(* Logix 5000 project; controller MV vendor 1 type 14 code 217 rev 31.11; software revision 31.00; part 22 of 53 *)
(* tags used below, declared in another part *)
   CheckTimeMask : INT;
   CWD : CHECKWORD_FLAGS;
   Delphi_Does_Eng_Func : BOOL;
   MC_CD_T1 : PlantItem;   // CD_T1
   MC_CD_T2 : PlantItem;   // CD_T2
   MC_CH2_LF1 : PlantItem;   // CH2_LF1
   MC_FL_D1 : PlantItem;   // FL_D1
   MC_FL_D2 : PlantItem;   // FL_D2
   MC_FL_PR : PlantItem;   // FL_PR
   MC_N255 : INT[255];   // CHECKWORDS Plant item checkword s
   MC_SPV1 : PlantItem;   // SPV1
   MC_SPV2 : PlantItem;   // SPV2
   MC_SPV3 : PlantItem;   // SPV3
   MC_SPV4 : PlantItem;   // SPV4
   MC_SPV5 : PlantItem;   // SPV5
   MC_SV1 : PlantItem;   // SV1
   MC_SV2 : PlantItem;   // SV2
   TempChecktime : DINT;
(* MC_Common, continued *)

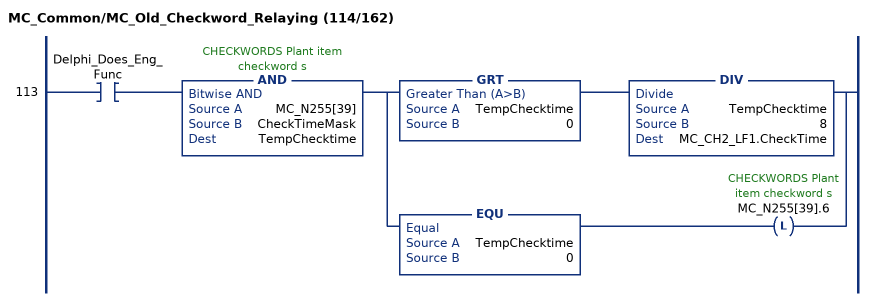
   [picture p386: MC_Common/MC_Old_Checkword_Relaying rungs 113-113]
   113: XIC(Delphi_Does_Eng_Func)AND(MC_N255[39],CheckTimeMask,TempChecktime)[GRT(TempChecktime,0) DIV(TempChecktime,8,MC_CH2_LF1.CheckTime) ,EQU(TempChecktime,0) OTL(MC_N255[39].6) ];
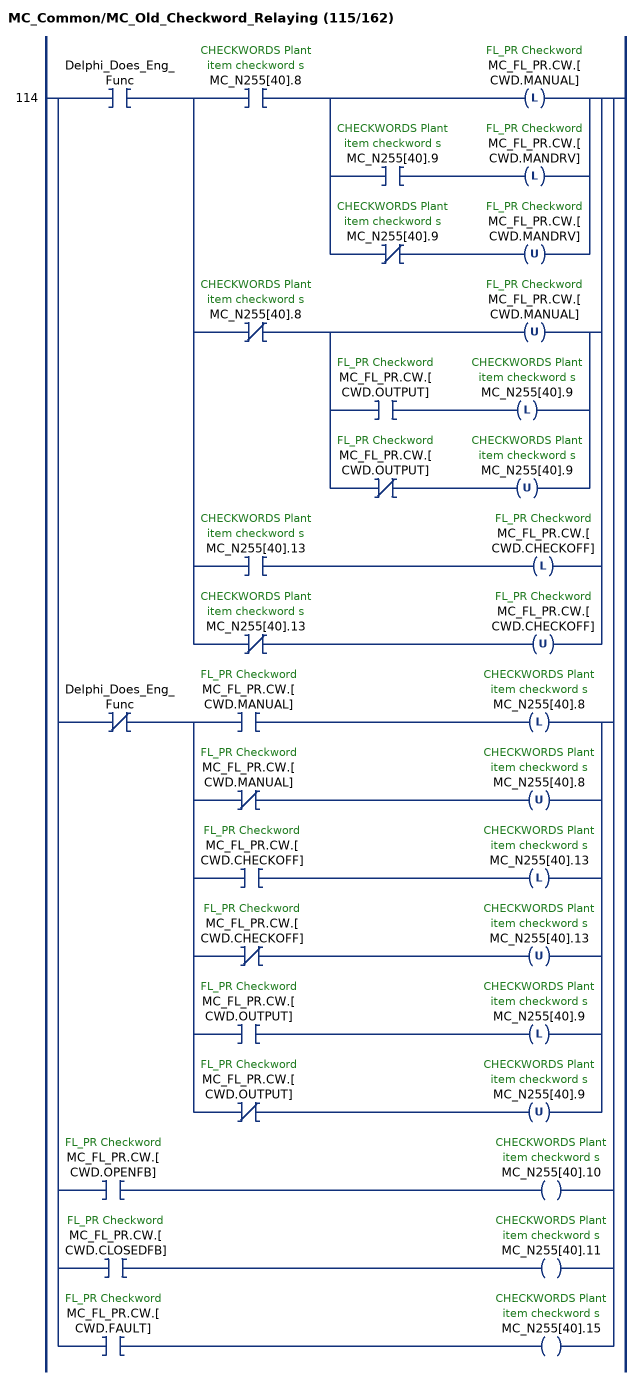
   114: [XIC(Delphi_Does_Eng_Func) [[XIC(MC_N255[40].8) [OTL(MC_FL_PR.CW.[CWD.MANUAL]) ,XIC(MC_N255[40].9) OTL(MC_FL_PR.CW.[CWD.MANDRV]) ,XIO(MC_N255[40].9) OTU(MC_FL_PR.CW.[CWD.MANDRV]) ] ,XIO(MC_N255[40].8) [OTU(MC_FL_PR.CW.[CWD.MANUAL]) ,[XIC(MC_FL_PR.CW.[CWD.OUTPUT]) OTL(MC_N255[40].9) ,XIO(MC_FL_PR.CW.[CWD.OUTPUT]) OTU(MC_N255[40].9) ] ] ] ,[XIC(MC_N255[40].13) OTL(MC_FL_PR.CW.[CWD.CHECKOFF]) ,XIO(MC_N255[40].13) OTU(MC_FL_PR.CW.[CWD.CHECKOFF]) ] ] ,XIO(Delphi_Does_Eng_Func) [[XIC(MC_FL_PR.CW.[CWD.MANUAL]) OTL(MC_N255[40].8) ,XIO(MC_FL_PR.CW.[CWD.MANUAL]) OTU(MC_N255[40].8) ] ,[XIC(MC_FL_PR.CW.[CWD.CHECKOFF]) OTL(MC_N255[40].13) ,XIO(MC_FL_PR.CW.[CWD.CHECKOFF]) OTU(MC_N255[40].13) ] ,[XIC(MC_FL_PR.CW.[CWD.OUTPUT]) OTL(MC_N255[40].9) ,XIO(MC_FL_PR.CW.[CWD.OUTPUT]) OTU(MC_N255[40].9) ] ] ,XIC(MC_FL_PR.CW.[CWD.OPENFB]) OTE(MC_N255[40].10) ,XIC(MC_FL_PR.CW.[CWD.CLOSEDFB]) OTE(MC_N255[40].11) ,XIC(MC_FL_PR.CW.[CWD.FAULT]) OTE(MC_N255[40].15) ];
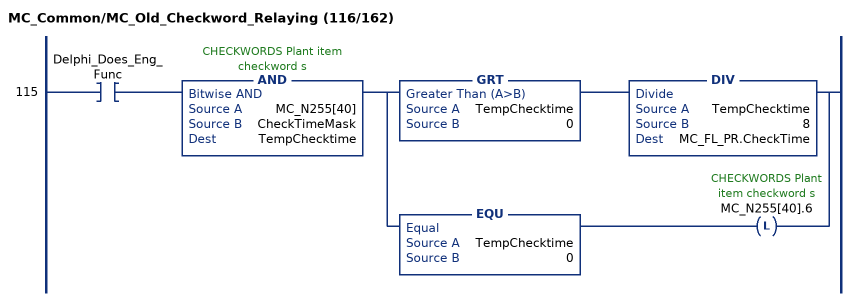
   115: XIC(Delphi_Does_Eng_Func)AND(MC_N255[40],CheckTimeMask,TempChecktime)[GRT(TempChecktime,0) DIV(TempChecktime,8,MC_FL_PR.CheckTime) ,EQU(TempChecktime,0) OTL(MC_N255[40].6) ];
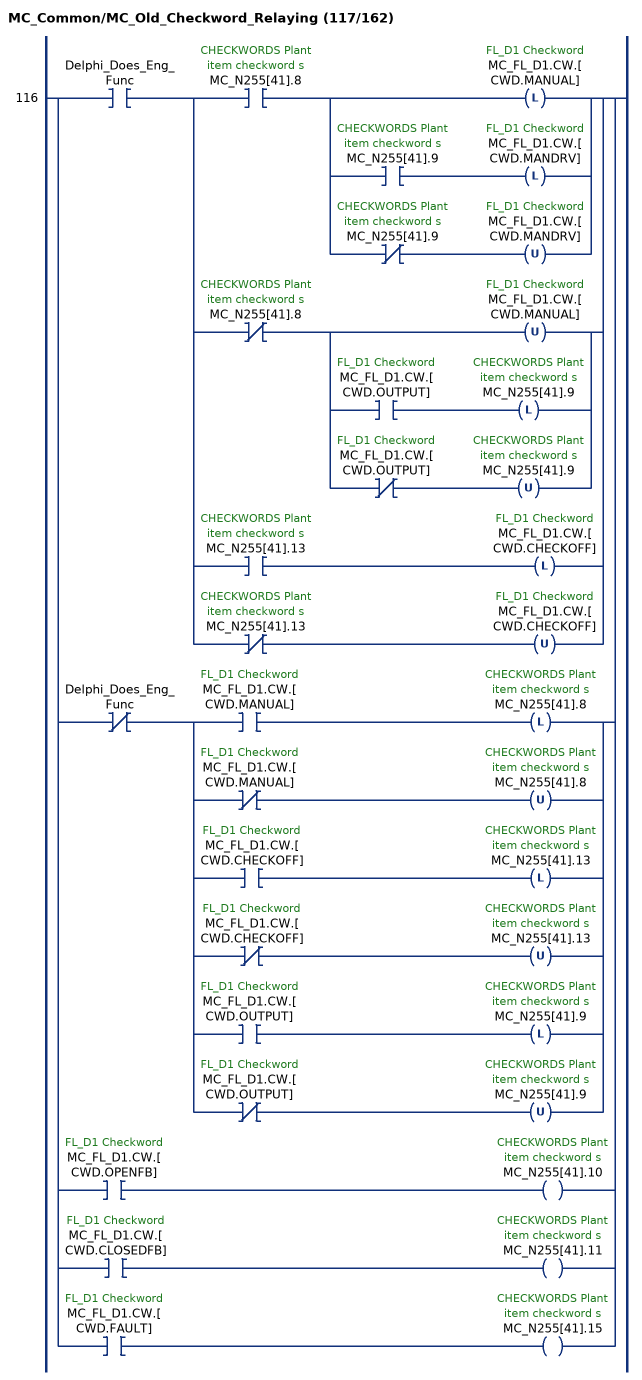
   116: [XIC(Delphi_Does_Eng_Func) [[XIC(MC_N255[41].8) [OTL(MC_FL_D1.CW.[CWD.MANUAL]) ,XIC(MC_N255[41].9) OTL(MC_FL_D1.CW.[CWD.MANDRV]) ,XIO(MC_N255[41].9) OTU(MC_FL_D1.CW.[CWD.MANDRV]) ] ,XIO(MC_N255[41].8) [OTU(MC_FL_D1.CW.[CWD.MANUAL]) ,[XIC(MC_FL_D1.CW.[CWD.OUTPUT]) OTL(MC_N255[41].9) ,XIO(MC_FL_D1.CW.[CWD.OUTPUT]) OTU(MC_N255[41].9) ] ] ] ,[XIC(MC_N255[41].13) OTL(MC_FL_D1.CW.[CWD.CHECKOFF]) ,XIO(MC_N255[41].13) OTU(MC_FL_D1.CW.[CWD.CHECKOFF]) ] ] ,XIO(Delphi_Does_Eng_Func) [[XIC(MC_FL_D1.CW.[CWD.MANUAL]) OTL(MC_N255[41].8) ,XIO(MC_FL_D1.CW.[CWD.MANUAL]) OTU(MC_N255[41].8) ] ,[XIC(MC_FL_D1.CW.[CWD.CHECKOFF]) OTL(MC_N255[41].13) ,XIO(MC_FL_D1.CW.[CWD.CHECKOFF]) OTU(MC_N255[41].13) ] ,[XIC(MC_FL_D1.CW.[CWD.OUTPUT]) OTL(MC_N255[41].9) ,XIO(MC_FL_D1.CW.[CWD.OUTPUT]) OTU(MC_N255[41].9) ] ] ,XIC(MC_FL_D1.CW.[CWD.OPENFB]) OTE(MC_N255[41].10) ,XIC(MC_FL_D1.CW.[CWD.CLOSEDFB]) OTE(MC_N255[41].11) ,XIC(MC_FL_D1.CW.[CWD.FAULT]) OTE(MC_N255[41].15) ];
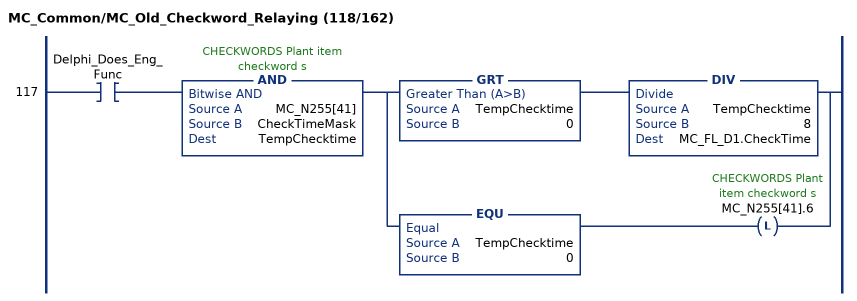
   117: XIC(Delphi_Does_Eng_Func)AND(MC_N255[41],CheckTimeMask,TempChecktime)[GRT(TempChecktime,0) DIV(TempChecktime,8,MC_FL_D1.CheckTime) ,EQU(TempChecktime,0) OTL(MC_N255[41].6) ];
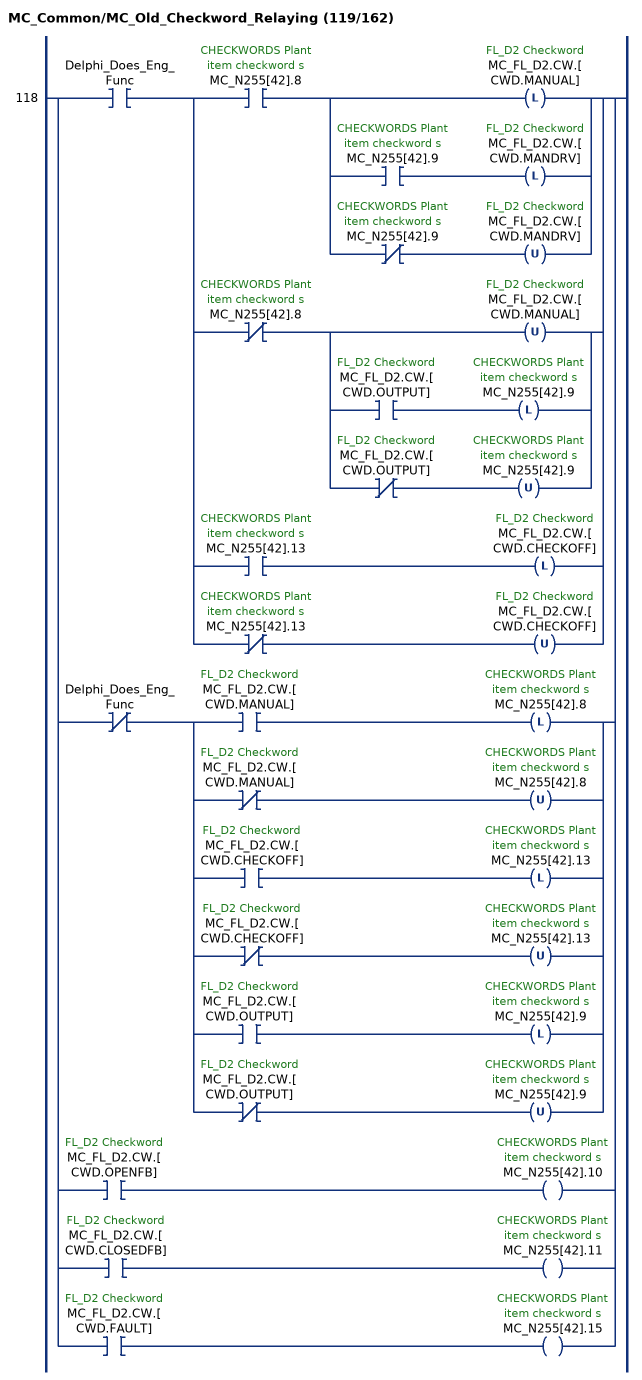
   118: [XIC(Delphi_Does_Eng_Func) [[XIC(MC_N255[42].8) [OTL(MC_FL_D2.CW.[CWD.MANUAL]) ,XIC(MC_N255[42].9) OTL(MC_FL_D2.CW.[CWD.MANDRV]) ,XIO(MC_N255[42].9) OTU(MC_FL_D2.CW.[CWD.MANDRV]) ] ,XIO(MC_N255[42].8) [OTU(MC_FL_D2.CW.[CWD.MANUAL]) ,[XIC(MC_FL_D2.CW.[CWD.OUTPUT]) OTL(MC_N255[42].9) ,XIO(MC_FL_D2.CW.[CWD.OUTPUT]) OTU(MC_N255[42].9) ] ] ] ,[XIC(MC_N255[42].13) OTL(MC_FL_D2.CW.[CWD.CHECKOFF]) ,XIO(MC_N255[42].13) OTU(MC_FL_D2.CW.[CWD.CHECKOFF]) ] ] ,XIO(Delphi_Does_Eng_Func) [[XIC(MC_FL_D2.CW.[CWD.MANUAL]) OTL(MC_N255[42].8) ,XIO(MC_FL_D2.CW.[CWD.MANUAL]) OTU(MC_N255[42].8) ] ,[XIC(MC_FL_D2.CW.[CWD.CHECKOFF]) OTL(MC_N255[42].13) ,XIO(MC_FL_D2.CW.[CWD.CHECKOFF]) OTU(MC_N255[42].13) ] ,[XIC(MC_FL_D2.CW.[CWD.OUTPUT]) OTL(MC_N255[42].9) ,XIO(MC_FL_D2.CW.[CWD.OUTPUT]) OTU(MC_N255[42].9) ] ] ,XIC(MC_FL_D2.CW.[CWD.OPENFB]) OTE(MC_N255[42].10) ,XIC(MC_FL_D2.CW.[CWD.CLOSEDFB]) OTE(MC_N255[42].11) ,XIC(MC_FL_D2.CW.[CWD.FAULT]) OTE(MC_N255[42].15) ];
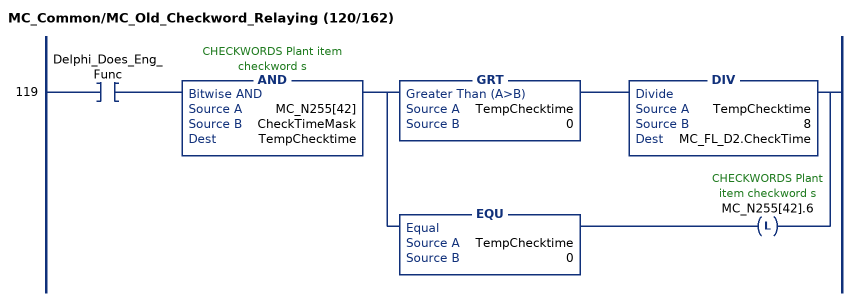
   119: XIC(Delphi_Does_Eng_Func)AND(MC_N255[42],CheckTimeMask,TempChecktime)[GRT(TempChecktime,0) DIV(TempChecktime,8,MC_FL_D2.CheckTime) ,EQU(TempChecktime,0) OTL(MC_N255[42].6) ];
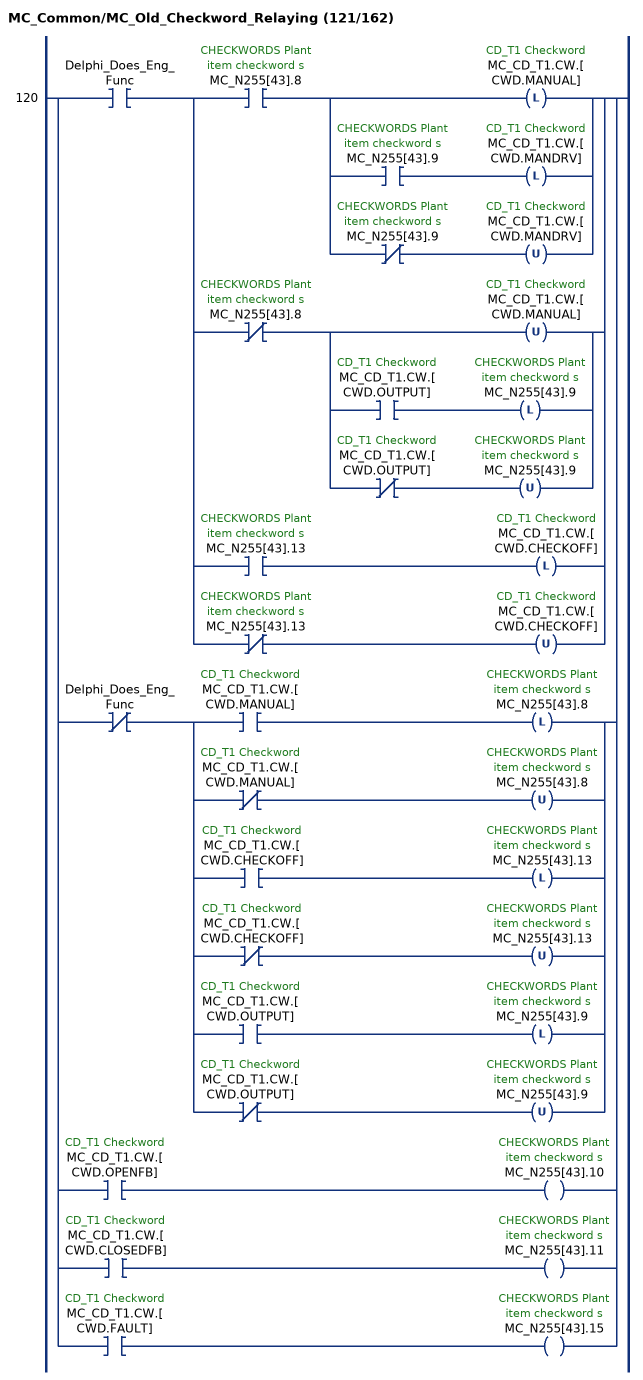
   120: [XIC(Delphi_Does_Eng_Func) [[XIC(MC_N255[43].8) [OTL(MC_CD_T1.CW.[CWD.MANUAL]) ,XIC(MC_N255[43].9) OTL(MC_CD_T1.CW.[CWD.MANDRV]) ,XIO(MC_N255[43].9) OTU(MC_CD_T1.CW.[CWD.MANDRV]) ] ,XIO(MC_N255[43].8) [OTU(MC_CD_T1.CW.[CWD.MANUAL]) ,[XIC(MC_CD_T1.CW.[CWD.OUTPUT]) OTL(MC_N255[43].9) ,XIO(MC_CD_T1.CW.[CWD.OUTPUT]) OTU(MC_N255[43].9) ] ] ] ,[XIC(MC_N255[43].13) OTL(MC_CD_T1.CW.[CWD.CHECKOFF]) ,XIO(MC_N255[43].13) OTU(MC_CD_T1.CW.[CWD.CHECKOFF]) ] ] ,XIO(Delphi_Does_Eng_Func) [[XIC(MC_CD_T1.CW.[CWD.MANUAL]) OTL(MC_N255[43].8) ,XIO(MC_CD_T1.CW.[CWD.MANUAL]) OTU(MC_N255[43].8) ] ,[XIC(MC_CD_T1.CW.[CWD.CHECKOFF]) OTL(MC_N255[43].13) ,XIO(MC_CD_T1.CW.[CWD.CHECKOFF]) OTU(MC_N255[43].13) ] ,[XIC(MC_CD_T1.CW.[CWD.OUTPUT]) OTL(MC_N255[43].9) ,XIO(MC_CD_T1.CW.[CWD.OUTPUT]) OTU(MC_N255[43].9) ] ] ,XIC(MC_CD_T1.CW.[CWD.OPENFB]) OTE(MC_N255[43].10) ,XIC(MC_CD_T1.CW.[CWD.CLOSEDFB]) OTE(MC_N255[43].11) ,XIC(MC_CD_T1.CW.[CWD.FAULT]) OTE(MC_N255[43].15) ];
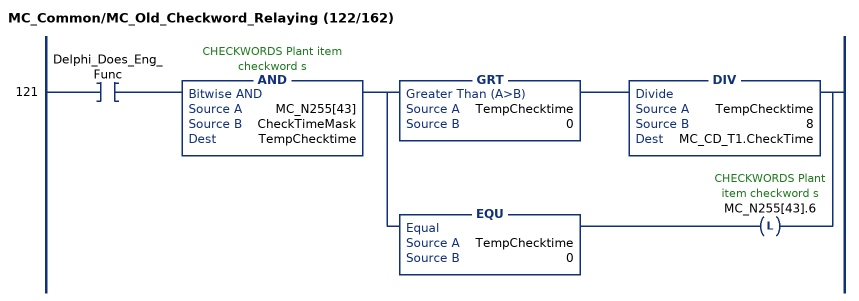
   121: XIC(Delphi_Does_Eng_Func)AND(MC_N255[43],CheckTimeMask,TempChecktime)[GRT(TempChecktime,0) DIV(TempChecktime,8,MC_CD_T1.CheckTime) ,EQU(TempChecktime,0) OTL(MC_N255[43].6) ];
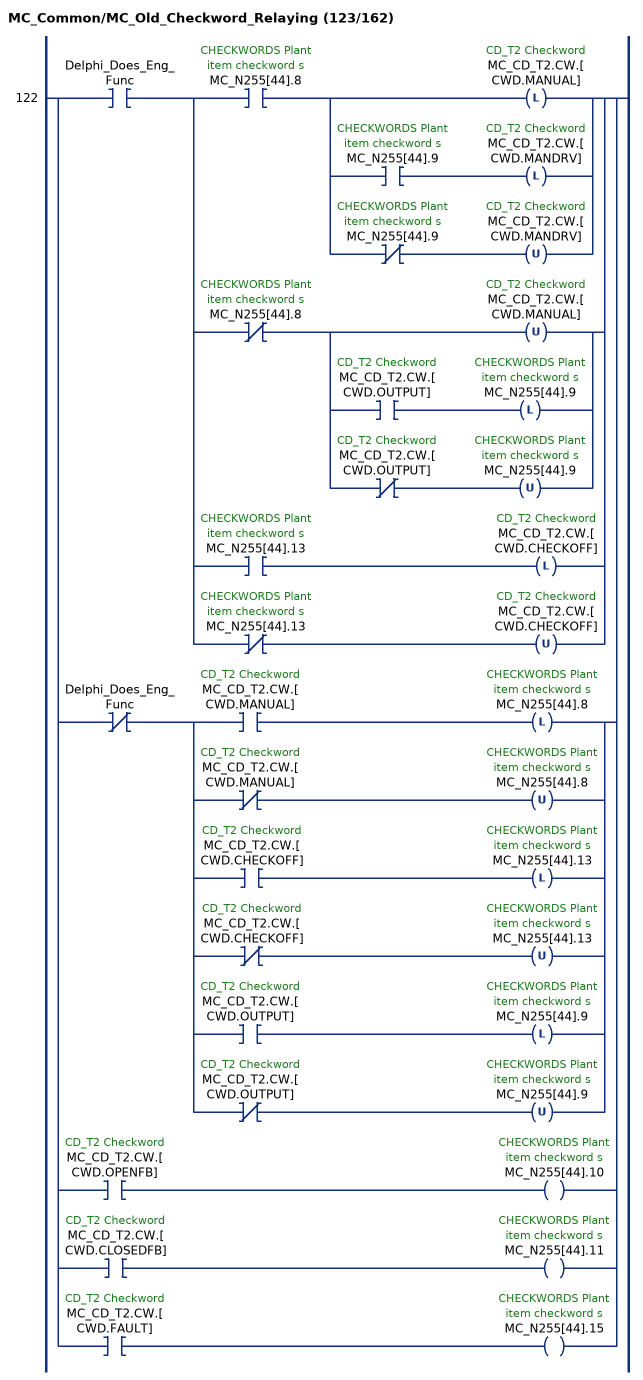
   122: [XIC(Delphi_Does_Eng_Func) [[XIC(MC_N255[44].8) [OTL(MC_CD_T2.CW.[CWD.MANUAL]) ,XIC(MC_N255[44].9) OTL(MC_CD_T2.CW.[CWD.MANDRV]) ,XIO(MC_N255[44].9) OTU(MC_CD_T2.CW.[CWD.MANDRV]) ] ,XIO(MC_N255[44].8) [OTU(MC_CD_T2.CW.[CWD.MANUAL]) ,[XIC(MC_CD_T2.CW.[CWD.OUTPUT]) OTL(MC_N255[44].9) ,XIO(MC_CD_T2.CW.[CWD.OUTPUT]) OTU(MC_N255[44].9) ] ] ] ,[XIC(MC_N255[44].13) OTL(MC_CD_T2.CW.[CWD.CHECKOFF]) ,XIO(MC_N255[44].13) OTU(MC_CD_T2.CW.[CWD.CHECKOFF]) ] ] ,XIO(Delphi_Does_Eng_Func) [[XIC(MC_CD_T2.CW.[CWD.MANUAL]) OTL(MC_N255[44].8) ,XIO(MC_CD_T2.CW.[CWD.MANUAL]) OTU(MC_N255[44].8) ] ,[XIC(MC_CD_T2.CW.[CWD.CHECKOFF]) OTL(MC_N255[44].13) ,XIO(MC_CD_T2.CW.[CWD.CHECKOFF]) OTU(MC_N255[44].13) ] ,[XIC(MC_CD_T2.CW.[CWD.OUTPUT]) OTL(MC_N255[44].9) ,XIO(MC_CD_T2.CW.[CWD.OUTPUT]) OTU(MC_N255[44].9) ] ] ,XIC(MC_CD_T2.CW.[CWD.OPENFB]) OTE(MC_N255[44].10) ,XIC(MC_CD_T2.CW.[CWD.CLOSEDFB]) OTE(MC_N255[44].11) ,XIC(MC_CD_T2.CW.[CWD.FAULT]) OTE(MC_N255[44].15) ];
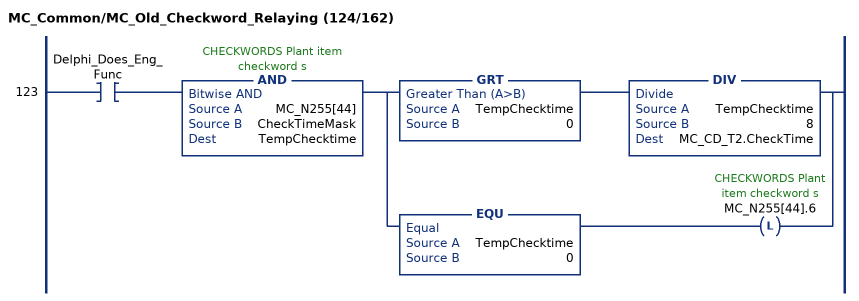
   123: XIC(Delphi_Does_Eng_Func)AND(MC_N255[44],CheckTimeMask,TempChecktime)[GRT(TempChecktime,0) DIV(TempChecktime,8,MC_CD_T2.CheckTime) ,EQU(TempChecktime,0) OTL(MC_N255[44].6) ];
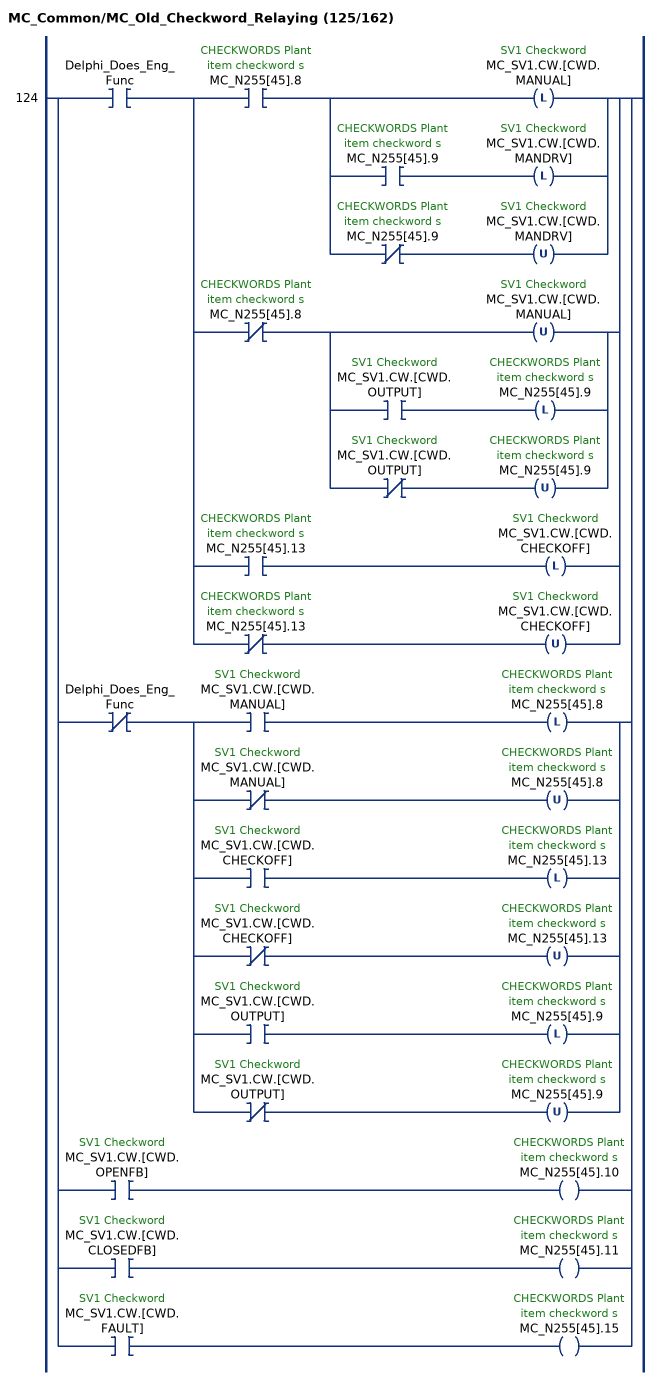
   124: [XIC(Delphi_Does_Eng_Func) [[XIC(MC_N255[45].8) [OTL(MC_SV1.CW.[CWD.MANUAL]) ,XIC(MC_N255[45].9) OTL(MC_SV1.CW.[CWD.MANDRV]) ,XIO(MC_N255[45].9) OTU(MC_SV1.CW.[CWD.MANDRV]) ] ,XIO(MC_N255[45].8) [OTU(MC_SV1.CW.[CWD.MANUAL]) ,[XIC(MC_SV1.CW.[CWD.OUTPUT]) OTL(MC_N255[45].9) ,XIO(MC_SV1.CW.[CWD.OUTPUT]) OTU(MC_N255[45].9) ] ] ] ,[XIC(MC_N255[45].13) OTL(MC_SV1.CW.[CWD.CHECKOFF]) ,XIO(MC_N255[45].13) OTU(MC_SV1.CW.[CWD.CHECKOFF]) ] ] ,XIO(Delphi_Does_Eng_Func) [[XIC(MC_SV1.CW.[CWD.MANUAL]) OTL(MC_N255[45].8) ,XIO(MC_SV1.CW.[CWD.MANUAL]) OTU(MC_N255[45].8) ] ,[XIC(MC_SV1.CW.[CWD.CHECKOFF]) OTL(MC_N255[45].13) ,XIO(MC_SV1.CW.[CWD.CHECKOFF]) OTU(MC_N255[45].13) ] ,[XIC(MC_SV1.CW.[CWD.OUTPUT]) OTL(MC_N255[45].9) ,XIO(MC_SV1.CW.[CWD.OUTPUT]) OTU(MC_N255[45].9) ] ] ,XIC(MC_SV1.CW.[CWD.OPENFB]) OTE(MC_N255[45].10) ,XIC(MC_SV1.CW.[CWD.CLOSEDFB]) OTE(MC_N255[45].11) ,XIC(MC_SV1.CW.[CWD.FAULT]) OTE(MC_N255[45].15) ];
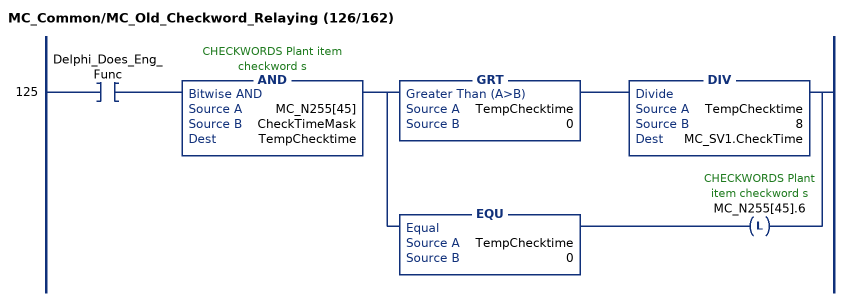
   125: XIC(Delphi_Does_Eng_Func)AND(MC_N255[45],CheckTimeMask,TempChecktime)[GRT(TempChecktime,0) DIV(TempChecktime,8,MC_SV1.CheckTime) ,EQU(TempChecktime,0) OTL(MC_N255[45].6) ];
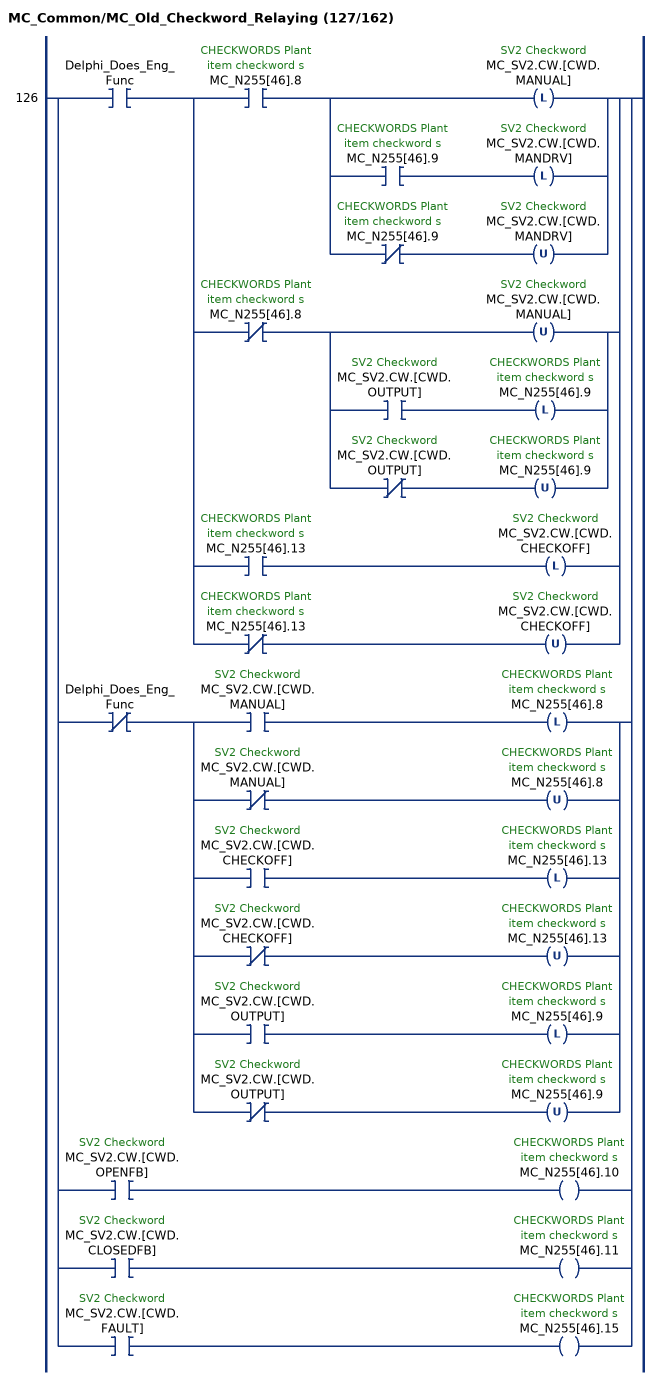
   126: [XIC(Delphi_Does_Eng_Func) [[XIC(MC_N255[46].8) [OTL(MC_SV2.CW.[CWD.MANUAL]) ,XIC(MC_N255[46].9) OTL(MC_SV2.CW.[CWD.MANDRV]) ,XIO(MC_N255[46].9) OTU(MC_SV2.CW.[CWD.MANDRV]) ] ,XIO(MC_N255[46].8) [OTU(MC_SV2.CW.[CWD.MANUAL]) ,[XIC(MC_SV2.CW.[CWD.OUTPUT]) OTL(MC_N255[46].9) ,XIO(MC_SV2.CW.[CWD.OUTPUT]) OTU(MC_N255[46].9) ] ] ] ,[XIC(MC_N255[46].13) OTL(MC_SV2.CW.[CWD.CHECKOFF]) ,XIO(MC_N255[46].13) OTU(MC_SV2.CW.[CWD.CHECKOFF]) ] ] ,XIO(Delphi_Does_Eng_Func) [[XIC(MC_SV2.CW.[CWD.MANUAL]) OTL(MC_N255[46].8) ,XIO(MC_SV2.CW.[CWD.MANUAL]) OTU(MC_N255[46].8) ] ,[XIC(MC_SV2.CW.[CWD.CHECKOFF]) OTL(MC_N255[46].13) ,XIO(MC_SV2.CW.[CWD.CHECKOFF]) OTU(MC_N255[46].13) ] ,[XIC(MC_SV2.CW.[CWD.OUTPUT]) OTL(MC_N255[46].9) ,XIO(MC_SV2.CW.[CWD.OUTPUT]) OTU(MC_N255[46].9) ] ] ,XIC(MC_SV2.CW.[CWD.OPENFB]) OTE(MC_N255[46].10) ,XIC(MC_SV2.CW.[CWD.CLOSEDFB]) OTE(MC_N255[46].11) ,XIC(MC_SV2.CW.[CWD.FAULT]) OTE(MC_N255[46].15) ];
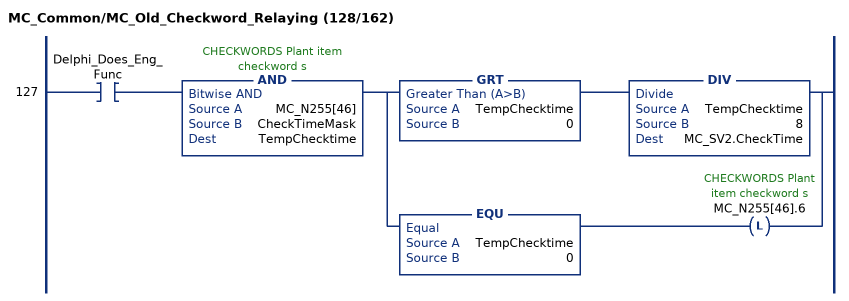
   127: XIC(Delphi_Does_Eng_Func)AND(MC_N255[46],CheckTimeMask,TempChecktime)[GRT(TempChecktime,0) DIV(TempChecktime,8,MC_SV2.CheckTime) ,EQU(TempChecktime,0) OTL(MC_N255[46].6) ];
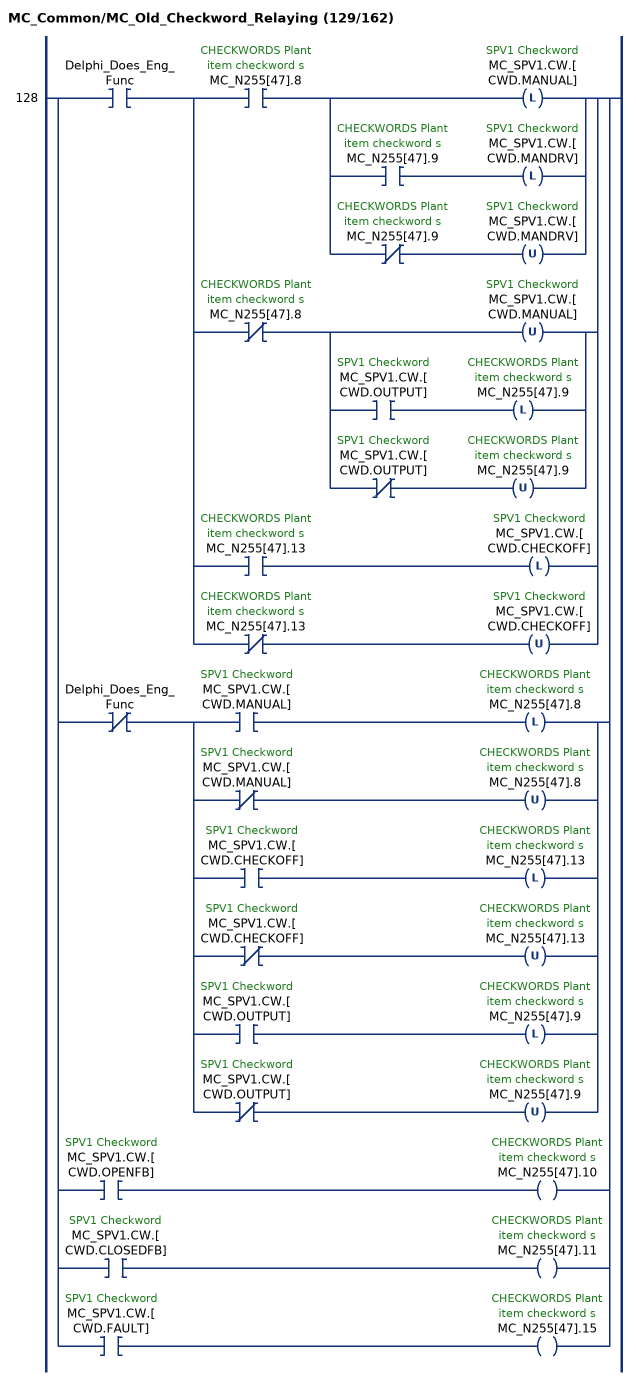
   128: [XIC(Delphi_Does_Eng_Func) [[XIC(MC_N255[47].8) [OTL(MC_SPV1.CW.[CWD.MANUAL]) ,XIC(MC_N255[47].9) OTL(MC_SPV1.CW.[CWD.MANDRV]) ,XIO(MC_N255[47].9) OTU(MC_SPV1.CW.[CWD.MANDRV]) ] ,XIO(MC_N255[47].8) [OTU(MC_SPV1.CW.[CWD.MANUAL]) ,[XIC(MC_SPV1.CW.[CWD.OUTPUT]) OTL(MC_N255[47].9) ,XIO(MC_SPV1.CW.[CWD.OUTPUT]) OTU(MC_N255[47].9) ] ] ] ,[XIC(MC_N255[47].13) OTL(MC_SPV1.CW.[CWD.CHECKOFF]) ,XIO(MC_N255[47].13) OTU(MC_SPV1.CW.[CWD.CHECKOFF]) ] ] ,XIO(Delphi_Does_Eng_Func) [[XIC(MC_SPV1.CW.[CWD.MANUAL]) OTL(MC_N255[47].8) ,XIO(MC_SPV1.CW.[CWD.MANUAL]) OTU(MC_N255[47].8) ] ,[XIC(MC_SPV1.CW.[CWD.CHECKOFF]) OTL(MC_N255[47].13) ,XIO(MC_SPV1.CW.[CWD.CHECKOFF]) OTU(MC_N255[47].13) ] ,[XIC(MC_SPV1.CW.[CWD.OUTPUT]) OTL(MC_N255[47].9) ,XIO(MC_SPV1.CW.[CWD.OUTPUT]) OTU(MC_N255[47].9) ] ] ,XIC(MC_SPV1.CW.[CWD.OPENFB]) OTE(MC_N255[47].10) ,XIC(MC_SPV1.CW.[CWD.CLOSEDFB]) OTE(MC_N255[47].11) ,XIC(MC_SPV1.CW.[CWD.FAULT]) OTE(MC_N255[47].15) ];
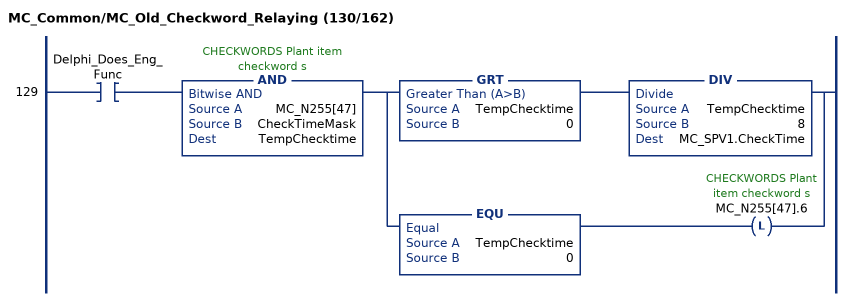
   129: XIC(Delphi_Does_Eng_Func)AND(MC_N255[47],CheckTimeMask,TempChecktime)[GRT(TempChecktime,0) DIV(TempChecktime,8,MC_SPV1.CheckTime) ,EQU(TempChecktime,0) OTL(MC_N255[47].6) ];
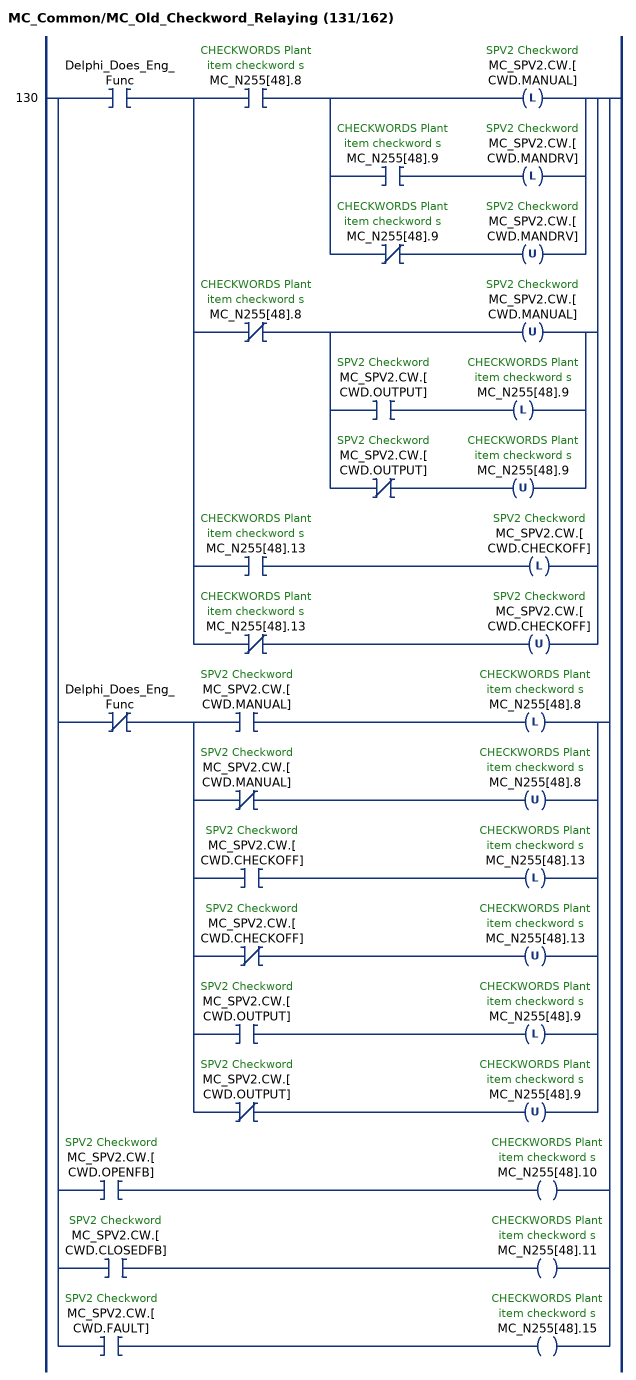
   130: [XIC(Delphi_Does_Eng_Func) [[XIC(MC_N255[48].8) [OTL(MC_SPV2.CW.[CWD.MANUAL]) ,XIC(MC_N255[48].9) OTL(MC_SPV2.CW.[CWD.MANDRV]) ,XIO(MC_N255[48].9) OTU(MC_SPV2.CW.[CWD.MANDRV]) ] ,XIO(MC_N255[48].8) [OTU(MC_SPV2.CW.[CWD.MANUAL]) ,[XIC(MC_SPV2.CW.[CWD.OUTPUT]) OTL(MC_N255[48].9) ,XIO(MC_SPV2.CW.[CWD.OUTPUT]) OTU(MC_N255[48].9) ] ] ] ,[XIC(MC_N255[48].13) OTL(MC_SPV2.CW.[CWD.CHECKOFF]) ,XIO(MC_N255[48].13) OTU(MC_SPV2.CW.[CWD.CHECKOFF]) ] ] ,XIO(Delphi_Does_Eng_Func) [[XIC(MC_SPV2.CW.[CWD.MANUAL]) OTL(MC_N255[48].8) ,XIO(MC_SPV2.CW.[CWD.MANUAL]) OTU(MC_N255[48].8) ] ,[XIC(MC_SPV2.CW.[CWD.CHECKOFF]) OTL(MC_N255[48].13) ,XIO(MC_SPV2.CW.[CWD.CHECKOFF]) OTU(MC_N255[48].13) ] ,[XIC(MC_SPV2.CW.[CWD.OUTPUT]) OTL(MC_N255[48].9) ,XIO(MC_SPV2.CW.[CWD.OUTPUT]) OTU(MC_N255[48].9) ] ] ,XIC(MC_SPV2.CW.[CWD.OPENFB]) OTE(MC_N255[48].10) ,XIC(MC_SPV2.CW.[CWD.CLOSEDFB]) OTE(MC_N255[48].11) ,XIC(MC_SPV2.CW.[CWD.FAULT]) OTE(MC_N255[48].15) ];
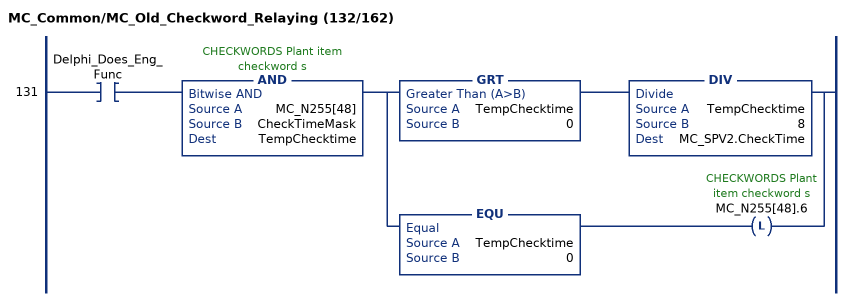
   131: XIC(Delphi_Does_Eng_Func)AND(MC_N255[48],CheckTimeMask,TempChecktime)[GRT(TempChecktime,0) DIV(TempChecktime,8,MC_SPV2.CheckTime) ,EQU(TempChecktime,0) OTL(MC_N255[48].6) ];
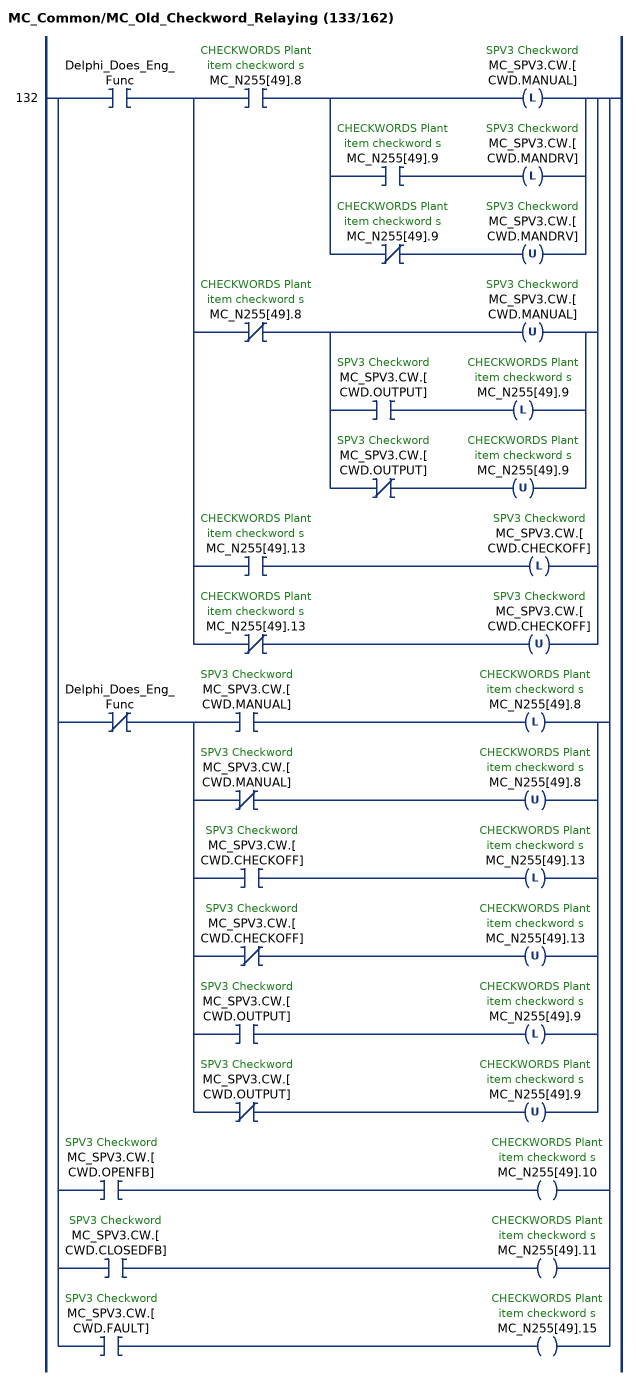
   132: [XIC(Delphi_Does_Eng_Func) [[XIC(MC_N255[49].8) [OTL(MC_SPV3.CW.[CWD.MANUAL]) ,XIC(MC_N255[49].9) OTL(MC_SPV3.CW.[CWD.MANDRV]) ,XIO(MC_N255[49].9) OTU(MC_SPV3.CW.[CWD.MANDRV]) ] ,XIO(MC_N255[49].8) [OTU(MC_SPV3.CW.[CWD.MANUAL]) ,[XIC(MC_SPV3.CW.[CWD.OUTPUT]) OTL(MC_N255[49].9) ,XIO(MC_SPV3.CW.[CWD.OUTPUT]) OTU(MC_N255[49].9) ] ] ] ,[XIC(MC_N255[49].13) OTL(MC_SPV3.CW.[CWD.CHECKOFF]) ,XIO(MC_N255[49].13) OTU(MC_SPV3.CW.[CWD.CHECKOFF]) ] ] ,XIO(Delphi_Does_Eng_Func) [[XIC(MC_SPV3.CW.[CWD.MANUAL]) OTL(MC_N255[49].8) ,XIO(MC_SPV3.CW.[CWD.MANUAL]) OTU(MC_N255[49].8) ] ,[XIC(MC_SPV3.CW.[CWD.CHECKOFF]) OTL(MC_N255[49].13) ,XIO(MC_SPV3.CW.[CWD.CHECKOFF]) OTU(MC_N255[49].13) ] ,[XIC(MC_SPV3.CW.[CWD.OUTPUT]) OTL(MC_N255[49].9) ,XIO(MC_SPV3.CW.[CWD.OUTPUT]) OTU(MC_N255[49].9) ] ] ,XIC(MC_SPV3.CW.[CWD.OPENFB]) OTE(MC_N255[49].10) ,XIC(MC_SPV3.CW.[CWD.CLOSEDFB]) OTE(MC_N255[49].11) ,XIC(MC_SPV3.CW.[CWD.FAULT]) OTE(MC_N255[49].15) ];
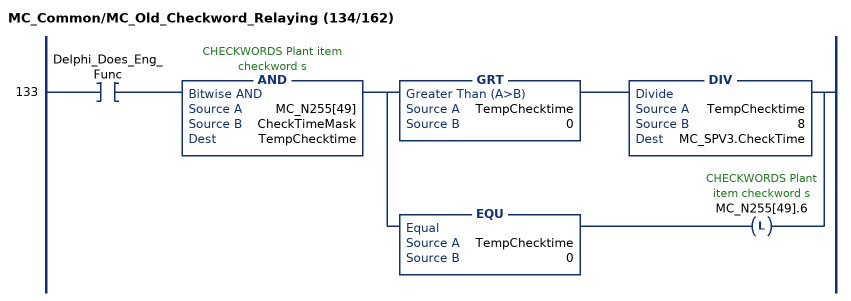
   133: XIC(Delphi_Does_Eng_Func)AND(MC_N255[49],CheckTimeMask,TempChecktime)[GRT(TempChecktime,0) DIV(TempChecktime,8,MC_SPV3.CheckTime) ,EQU(TempChecktime,0) OTL(MC_N255[49].6) ];
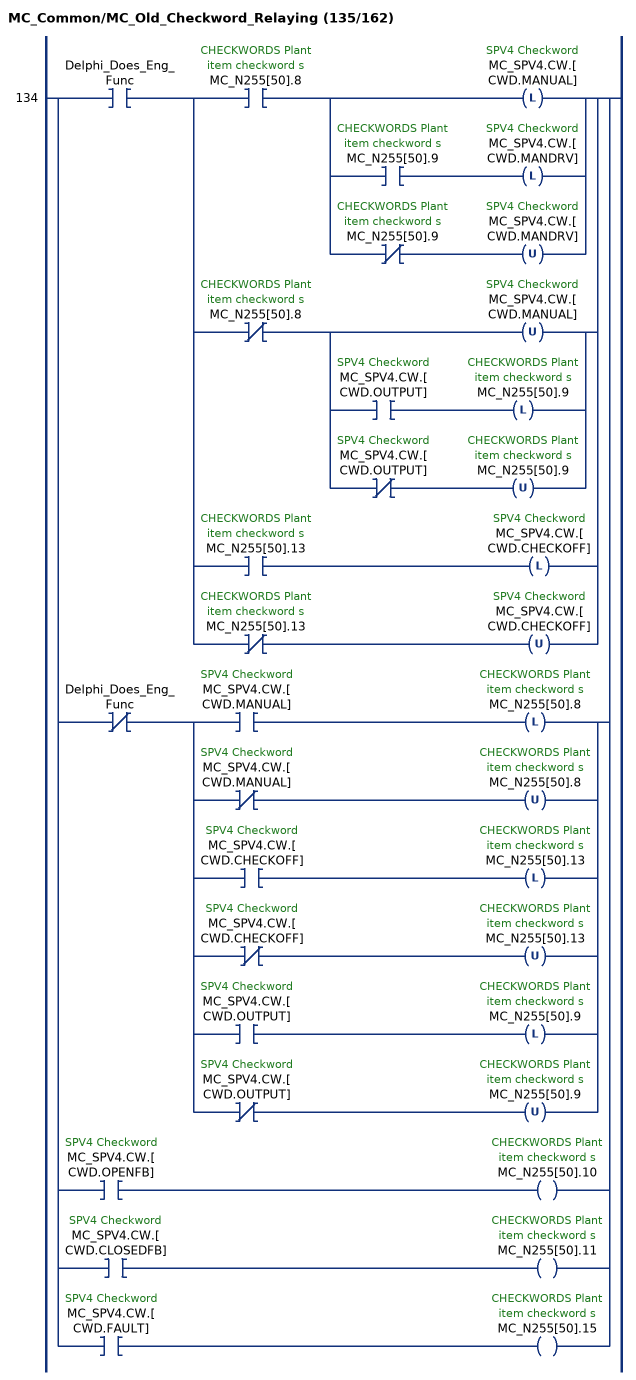
   134: [XIC(Delphi_Does_Eng_Func) [[XIC(MC_N255[50].8) [OTL(MC_SPV4.CW.[CWD.MANUAL]) ,XIC(MC_N255[50].9) OTL(MC_SPV4.CW.[CWD.MANDRV]) ,XIO(MC_N255[50].9) OTU(MC_SPV4.CW.[CWD.MANDRV]) ] ,XIO(MC_N255[50].8) [OTU(MC_SPV4.CW.[CWD.MANUAL]) ,[XIC(MC_SPV4.CW.[CWD.OUTPUT]) OTL(MC_N255[50].9) ,XIO(MC_SPV4.CW.[CWD.OUTPUT]) OTU(MC_N255[50].9) ] ] ] ,[XIC(MC_N255[50].13) OTL(MC_SPV4.CW.[CWD.CHECKOFF]) ,XIO(MC_N255[50].13) OTU(MC_SPV4.CW.[CWD.CHECKOFF]) ] ] ,XIO(Delphi_Does_Eng_Func) [[XIC(MC_SPV4.CW.[CWD.MANUAL]) OTL(MC_N255[50].8) ,XIO(MC_SPV4.CW.[CWD.MANUAL]) OTU(MC_N255[50].8) ] ,[XIC(MC_SPV4.CW.[CWD.CHECKOFF]) OTL(MC_N255[50].13) ,XIO(MC_SPV4.CW.[CWD.CHECKOFF]) OTU(MC_N255[50].13) ] ,[XIC(MC_SPV4.CW.[CWD.OUTPUT]) OTL(MC_N255[50].9) ,XIO(MC_SPV4.CW.[CWD.OUTPUT]) OTU(MC_N255[50].9) ] ] ,XIC(MC_SPV4.CW.[CWD.OPENFB]) OTE(MC_N255[50].10) ,XIC(MC_SPV4.CW.[CWD.CLOSEDFB]) OTE(MC_N255[50].11) ,XIC(MC_SPV4.CW.[CWD.FAULT]) OTE(MC_N255[50].15) ];
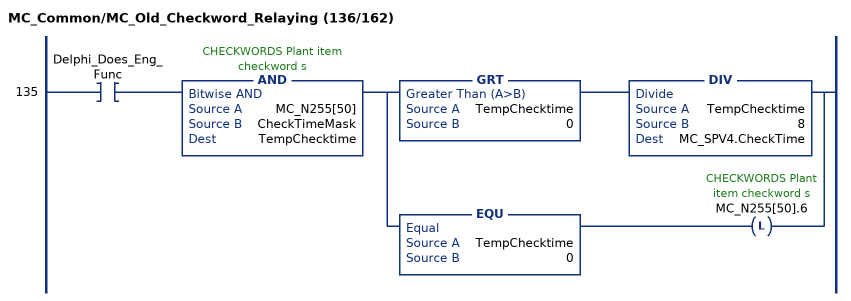
   135: XIC(Delphi_Does_Eng_Func)AND(MC_N255[50],CheckTimeMask,TempChecktime)[GRT(TempChecktime,0) DIV(TempChecktime,8,MC_SPV4.CheckTime) ,EQU(TempChecktime,0) OTL(MC_N255[50].6) ];
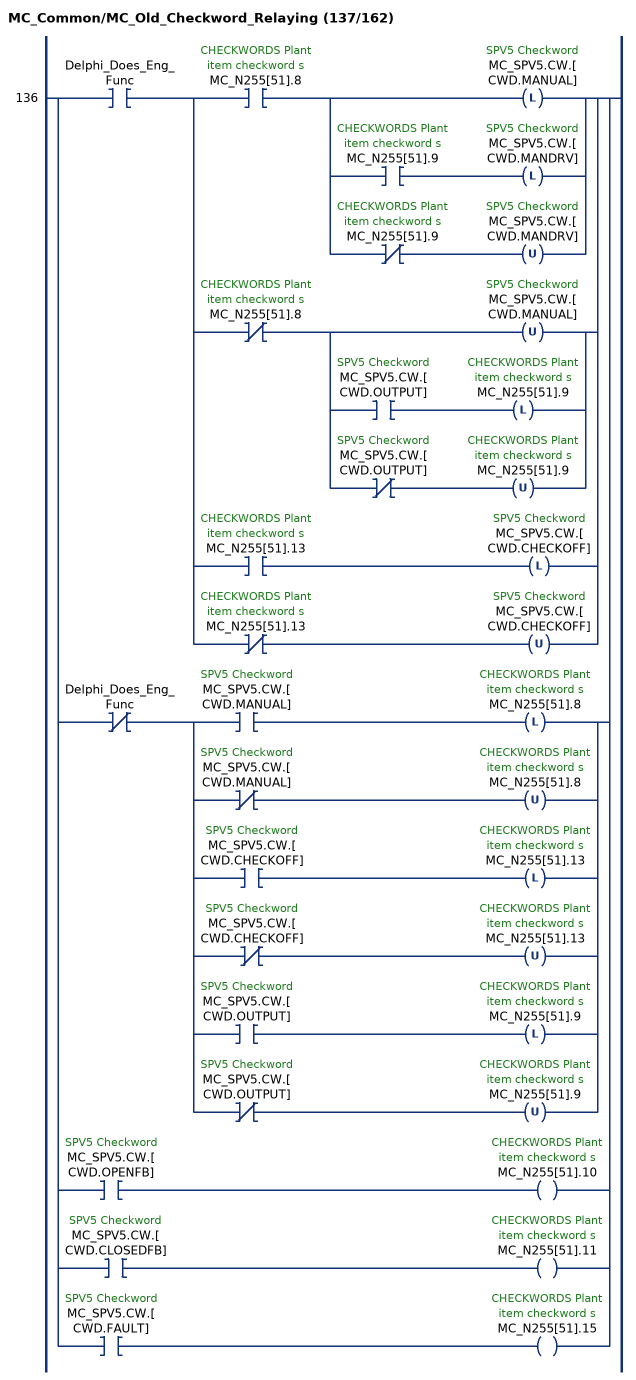
   136: [XIC(Delphi_Does_Eng_Func) [[XIC(MC_N255[51].8) [OTL(MC_SPV5.CW.[CWD.MANUAL]) ,XIC(MC_N255[51].9) OTL(MC_SPV5.CW.[CWD.MANDRV]) ,XIO(MC_N255[51].9) OTU(MC_SPV5.CW.[CWD.MANDRV]) ] ,XIO(MC_N255[51].8) [OTU(MC_SPV5.CW.[CWD.MANUAL]) ,[XIC(MC_SPV5.CW.[CWD.OUTPUT]) OTL(MC_N255[51].9) ,XIO(MC_SPV5.CW.[CWD.OUTPUT]) OTU(MC_N255[51].9) ] ] ] ,[XIC(MC_N255[51].13) OTL(MC_SPV5.CW.[CWD.CHECKOFF]) ,XIO(MC_N255[51].13) OTU(MC_SPV5.CW.[CWD.CHECKOFF]) ] ] ,XIO(Delphi_Does_Eng_Func) [[XIC(MC_SPV5.CW.[CWD.MANUAL]) OTL(MC_N255[51].8) ,XIO(MC_SPV5.CW.[CWD.MANUAL]) OTU(MC_N255[51].8) ] ,[XIC(MC_SPV5.CW.[CWD.CHECKOFF]) OTL(MC_N255[51].13) ,XIO(MC_SPV5.CW.[CWD.CHECKOFF]) OTU(MC_N255[51].13) ] ,[XIC(MC_SPV5.CW.[CWD.OUTPUT]) OTL(MC_N255[51].9) ,XIO(MC_SPV5.CW.[CWD.OUTPUT]) OTU(MC_N255[51].9) ] ] ,XIC(MC_SPV5.CW.[CWD.OPENFB]) OTE(MC_N255[51].10) ,XIC(MC_SPV5.CW.[CWD.CLOSEDFB]) OTE(MC_N255[51].11) ,XIC(MC_SPV5.CW.[CWD.FAULT]) OTE(MC_N255[51].15) ];
